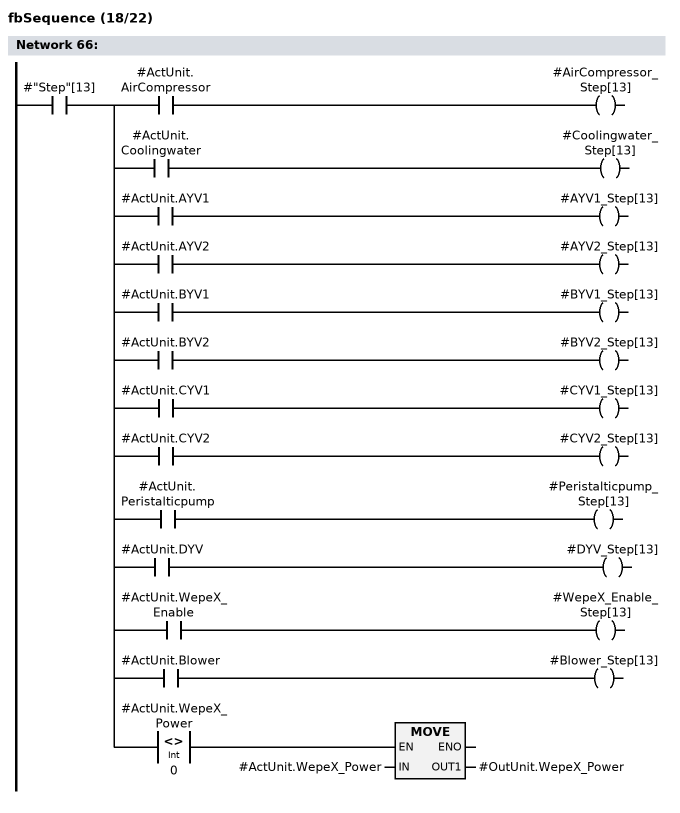
   RUNG wire#powerrail
      Contact( #"Step"[13] )
      wire#w1
      Contact( #ActUnit.AirCompressor )
      Coil( #AirCompressor_Step[13] )
   END_RUNG
   RUNG wire#w1
      Contact( #ActUnit.Coolingwater )
      Coil( #Coolingwater_Step[13] )
   END_RUNG
   RUNG wire#w1
      Contact( #ActUnit.AYV1 )
      Coil( #AYV1_Step[13] )
   END_RUNG
   RUNG wire#w1
      Contact( #ActUnit.AYV2 )
      Coil( #AYV2_Step[13] )
   END_RUNG
   RUNG wire#w1
      Contact( #ActUnit.BYV1 )
      Coil( #BYV1_Step[13] )
   END_RUNG
   RUNG wire#w1
      Contact( #ActUnit.BYV2 )
      Coil( #BYV2_Step[13] )
   END_RUNG
   RUNG wire#w1
      Contact( #ActUnit.CYV1 )
      Coil( #CYV1_Step[13] )
   END_RUNG
   RUNG wire#w1
      Contact( #ActUnit.CYV2 )
      Coil( #CYV2_Step[13] )
   END_RUNG
   RUNG wire#w1
      Contact( #ActUnit.Peristalticpump )
      Coil( #Peristalticpump_Step[13] )
   END_RUNG
   RUNG wire#w1
      Contact( #ActUnit.DYV )
      Coil( #DYV_Step[13] )
   END_RUNG
   RUNG wire#w1
      Contact( #ActUnit.WepeX_Enable )
      Coil( #WepeX_Enable_Step[13] )
   END_RUNG
   RUNG wire#w1
      Contact( #ActUnit.Blower )
      Coil( #Blower_Step[13] )
   END_RUNG
   RUNG wire#w1
      { S7_Templates := "SrcType := Int" } NE_Contact(in1 := #ActUnit.WepeX_Power, in2 := 0)
      Move(in := #ActUnit.WepeX_Power, out1 => #OutUnit.WepeX_Power)
   END_RUNG
   // the same network as SCL:
   #AirCompressor_Step[13] := #"Step"[13] AND #ActUnit.AirCompressor;
   #Coolingwater_Step[13] := #"Step"[13] AND #ActUnit.Coolingwater;
   #AYV1_Step[13] := #"Step"[13] AND #ActUnit.AYV1;
   #AYV2_Step[13] := #"Step"[13] AND #ActUnit.AYV2;
   #BYV1_Step[13] := #"Step"[13] AND #ActUnit.BYV1;
   #BYV2_Step[13] := #"Step"[13] AND #ActUnit.BYV2;
   #CYV1_Step[13] := #"Step"[13] AND #ActUnit.CYV1;
   #CYV2_Step[13] := #"Step"[13] AND #ActUnit.CYV2;
   #Peristalticpump_Step[13] := #"Step"[13] AND #ActUnit.Peristalticpump;
   #DYV_Step[13] := #"Step"[13] AND #ActUnit.DYV;
   #WepeX_Enable_Step[13] := #"Step"[13] AND #ActUnit.WepeX_Enable;
   #Blower_Step[13] := #"Step"[13] AND #ActUnit.Blower;
   IF #"Step"[13] AND (#ActUnit.WepeX_Power <> 0) THEN #OutUnit.WepeX_Power := #ActUnit.WepeX_Power; END_IF;
END_REGION

REGION Network 67
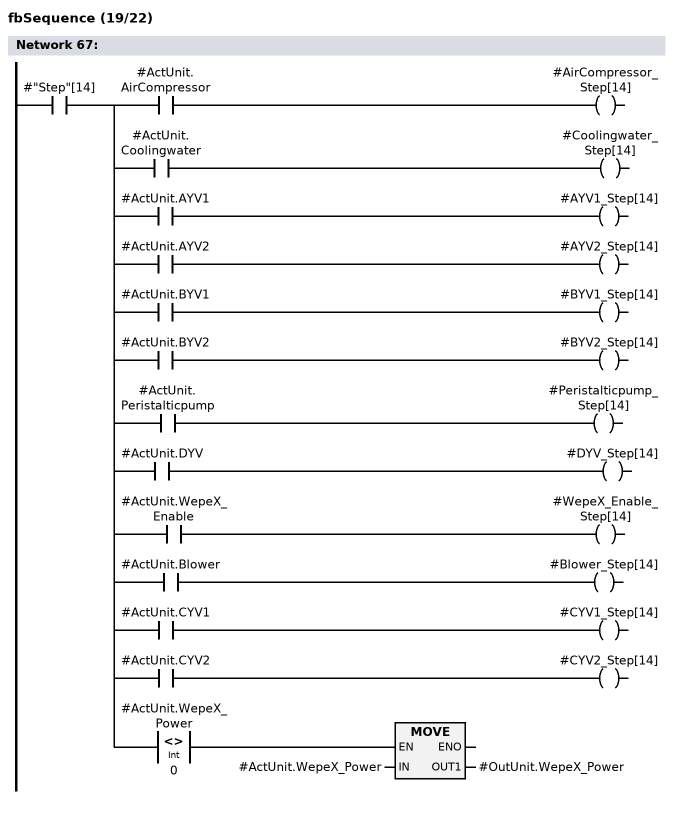
   RUNG wire#powerrail
      Contact( #"Step"[14] )
      wire#w1
      Contact( #ActUnit.AirCompressor )
      Coil( #AirCompressor_Step[14] )
   END_RUNG
   RUNG wire#w1
      Contact( #ActUnit.Coolingwater )
      Coil( #Coolingwater_Step[14] )
   END_RUNG
   RUNG wire#w1
      Contact( #ActUnit.AYV1 )
      Coil( #AYV1_Step[14] )
   END_RUNG
   RUNG wire#w1
      Contact( #ActUnit.AYV2 )
      Coil( #AYV2_Step[14] )
   END_RUNG
   RUNG wire#w1
      Contact( #ActUnit.BYV1 )
      Coil( #BYV1_Step[14] )
   END_RUNG
   RUNG wire#w1
      Contact( #ActUnit.BYV2 )
      Coil( #BYV2_Step[14] )
   END_RUNG
   RUNG wire#w1
      Contact( #ActUnit.Peristalticpump )
      Coil( #Peristalticpump_Step[14] )
   END_RUNG
   RUNG wire#w1
      Contact( #ActUnit.DYV )
      Coil( #DYV_Step[14] )
   END_RUNG
   RUNG wire#w1
      Contact( #ActUnit.WepeX_Enable )
      Coil( #WepeX_Enable_Step[14] )
   END_RUNG
   RUNG wire#w1
      Contact( #ActUnit.Blower )
      Coil( #Blower_Step[14] )
   END_RUNG
   RUNG wire#w1
      Contact( #ActUnit.CYV1 )
      Coil( #CYV1_Step[14] )
   END_RUNG
   RUNG wire#w1
      Contact( #ActUnit.CYV2 )
      Coil( #CYV2_Step[14] )
   END_RUNG
   RUNG wire#w1
      { S7_Templates := "SrcType := Int" } NE_Contact(in1 := #ActUnit.WepeX_Power, in2 := 0)
      Move(in := #ActUnit.WepeX_Power, out1 => #OutUnit.WepeX_Power)
   END_RUNG
   // the same network as SCL:
   #AirCompressor_Step[14] := #"Step"[14] AND #ActUnit.AirCompressor;
   #Coolingwater_Step[14] := #"Step"[14] AND #ActUnit.Coolingwater;
   #AYV1_Step[14] := #"Step"[14] AND #ActUnit.AYV1;
   #AYV2_Step[14] := #"Step"[14] AND #ActUnit.AYV2;
   #BYV1_Step[14] := #"Step"[14] AND #ActUnit.BYV1;
   #BYV2_Step[14] := #"Step"[14] AND #ActUnit.BYV2;
   #Peristalticpump_Step[14] := #"Step"[14] AND #ActUnit.Peristalticpump;
   #DYV_Step[14] := #"Step"[14] AND #ActUnit.DYV;
   #WepeX_Enable_Step[14] := #"Step"[14] AND #ActUnit.WepeX_Enable;
   #Blower_Step[14] := #"Step"[14] AND #ActUnit.Blower;
   #CYV1_Step[14] := #"Step"[14] AND #ActUnit.CYV1;
   #CYV2_Step[14] := #"Step"[14] AND #ActUnit.CYV2;
   IF #"Step"[14] AND (#ActUnit.WepeX_Power <> 0) THEN #OutUnit.WepeX_Power := #ActUnit.WepeX_Power; END_IF;
END_REGION

REGION Network 68
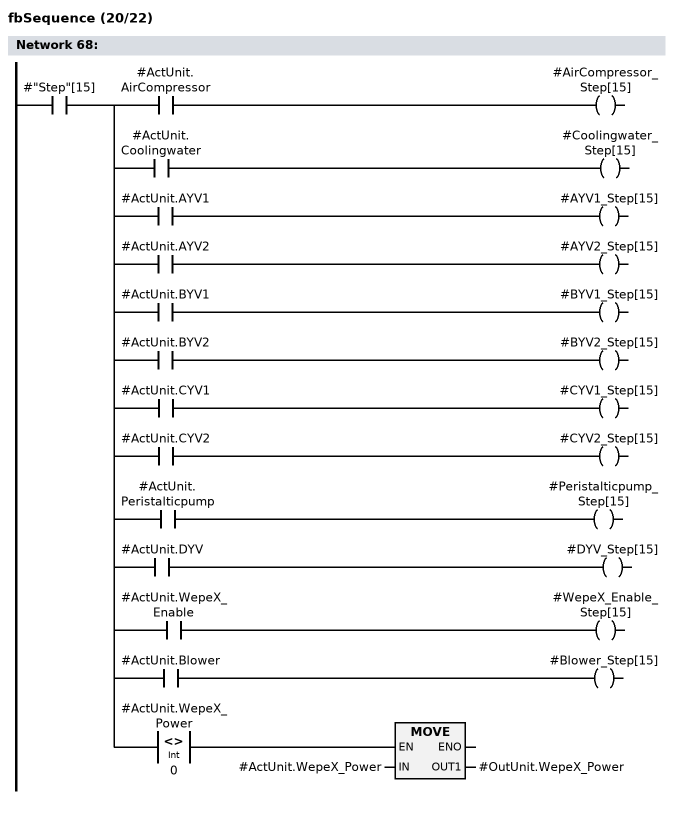
   RUNG wire#powerrail
      Contact( #"Step"[15] )
      wire#w1
      Contact( #ActUnit.AirCompressor )
      Coil( #AirCompressor_Step[15] )
   END_RUNG
   RUNG wire#w1
      Contact( #ActUnit.Coolingwater )
      Coil( #Coolingwater_Step[15] )
   END_RUNG
   RUNG wire#w1
      Contact( #ActUnit.AYV1 )
      Coil( #AYV1_Step[15] )
   END_RUNG
   RUNG wire#w1
      Contact( #ActUnit.AYV2 )
      Coil( #AYV2_Step[15] )
   END_RUNG
   RUNG wire#w1
      Contact( #ActUnit.BYV1 )
      Coil( #BYV1_Step[15] )
   END_RUNG
   RUNG wire#w1
      Contact( #ActUnit.BYV2 )
      Coil( #BYV2_Step[15] )
   END_RUNG
   RUNG wire#w1
      Contact( #ActUnit.CYV1 )
      Coil( #CYV1_Step[15] )
   END_RUNG
   RUNG wire#w1
      Contact( #ActUnit.CYV2 )
      Coil( #CYV2_Step[15] )
   END_RUNG
   RUNG wire#w1
      Contact( #ActUnit.Peristalticpump )
      Coil( #Peristalticpump_Step[15] )
   END_RUNG
   RUNG wire#w1
      Contact( #ActUnit.DYV )
      Coil( #DYV_Step[15] )
   END_RUNG
   RUNG wire#w1
      Contact( #ActUnit.WepeX_Enable )
      Coil( #WepeX_Enable_Step[15] )
   END_RUNG
   RUNG wire#w1
      Contact( #ActUnit.Blower )
      Coil( #Blower_Step[15] )
   END_RUNG
   RUNG wire#w1
      { S7_Templates := "SrcType := Int" } NE_Contact(in1 := #ActUnit.WepeX_Power, in2 := 0)
      Move(in := #ActUnit.WepeX_Power, out1 => #OutUnit.WepeX_Power)
   END_RUNG
   // the same network as SCL:
   #AirCompressor_Step[15] := #"Step"[15] AND #ActUnit.AirCompressor;
   #Coolingwater_Step[15] := #"Step"[15] AND #ActUnit.Coolingwater;
   #AYV1_Step[15] := #"Step"[15] AND #ActUnit.AYV1;
   #AYV2_Step[15] := #"Step"[15] AND #ActUnit.AYV2;
   #BYV1_Step[15] := #"Step"[15] AND #ActUnit.BYV1;
   #BYV2_Step[15] := #"Step"[15] AND #ActUnit.BYV2;
   #CYV1_Step[15] := #"Step"[15] AND #ActUnit.CYV1;
   #CYV2_Step[15] := #"Step"[15] AND #ActUnit.CYV2;
   #Peristalticpump_Step[15] := #"Step"[15] AND #ActUnit.Peristalticpump;
   #DYV_Step[15] := #"Step"[15] AND #ActUnit.DYV;
   #WepeX_Enable_Step[15] := #"Step"[15] AND #ActUnit.WepeX_Enable;
   #Blower_Step[15] := #"Step"[15] AND #ActUnit.Blower;
   IF #"Step"[15] AND (#ActUnit.WepeX_Power <> 0) THEN #OutUnit.WepeX_Power := #ActUnit.WepeX_Power; END_IF;
END_REGION

REGION Network 69
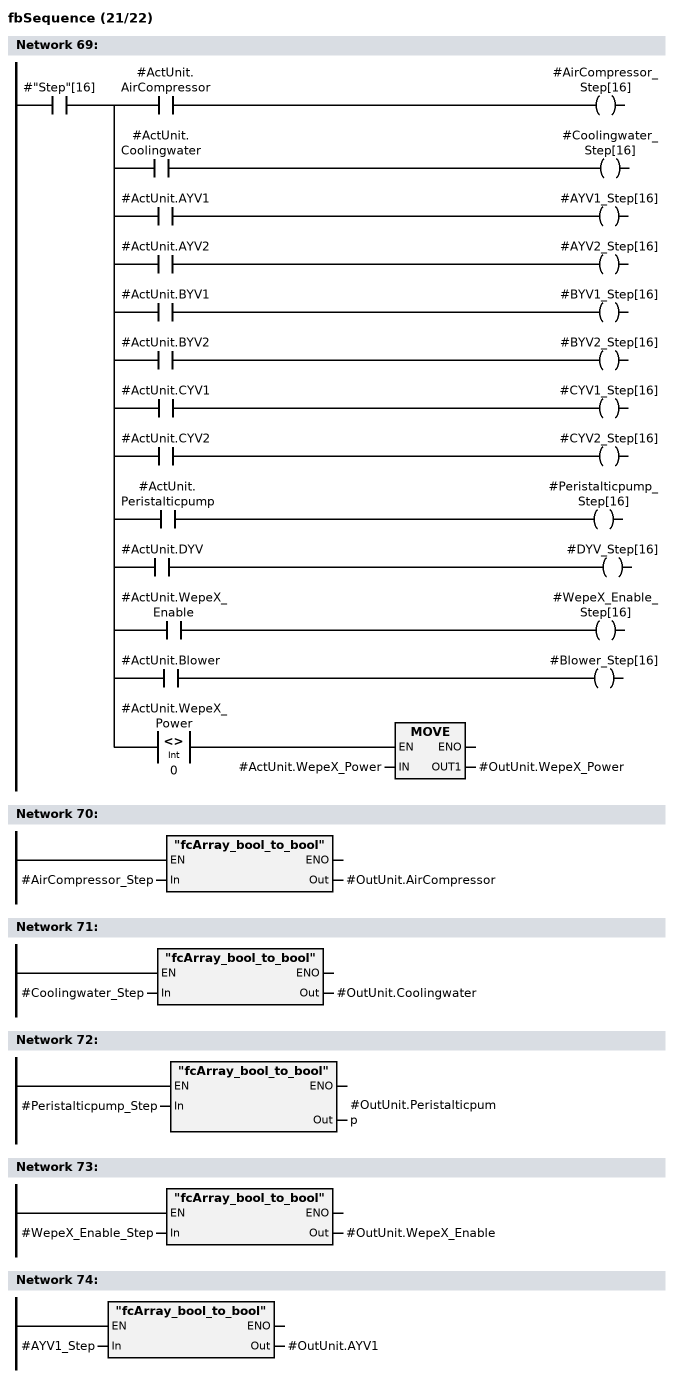
   RUNG wire#powerrail
      Contact( #"Step"[16] )
      wire#w1
      Contact( #ActUnit.AirCompressor )
      Coil( #AirCompressor_Step[16] )
   END_RUNG
   RUNG wire#w1
      Contact( #ActUnit.Coolingwater )
      Coil( #Coolingwater_Step[16] )
   END_RUNG
   RUNG wire#w1
      Contact( #ActUnit.AYV1 )
      Coil( #AYV1_Step[16] )
   END_RUNG
   RUNG wire#w1
      Contact( #ActUnit.AYV2 )
      Coil( #AYV2_Step[16] )
   END_RUNG
   RUNG wire#w1
      Contact( #ActUnit.BYV1 )
      Coil( #BYV1_Step[16] )
   END_RUNG
   RUNG wire#w1
      Contact( #ActUnit.BYV2 )
      Coil( #BYV2_Step[16] )
   END_RUNG
   RUNG wire#w1
      Contact( #ActUnit.CYV1 )
      Coil( #CYV1_Step[16] )
   END_RUNG
   RUNG wire#w1
      Contact( #ActUnit.CYV2 )
      Coil( #CYV2_Step[16] )
   END_RUNG
   RUNG wire#w1
      Contact( #ActUnit.Peristalticpump )
      Coil( #Peristalticpump_Step[16] )
   END_RUNG
   RUNG wire#w1
      Contact( #ActUnit.DYV )
      Coil( #DYV_Step[16] )
   END_RUNG
   RUNG wire#w1
      Contact( #ActUnit.WepeX_Enable )
      Coil( #WepeX_Enable_Step[16] )
   END_RUNG
   RUNG wire#w1
      Contact( #ActUnit.Blower )
      Coil( #Blower_Step[16] )
   END_RUNG
   RUNG wire#w1
      { S7_Templates := "SrcType := Int" } NE_Contact(in1 := #ActUnit.WepeX_Power, in2 := 0)
      Move(in := #ActUnit.WepeX_Power, out1 => #OutUnit.WepeX_Power)
   END_RUNG
   // the same network as SCL:
   #AirCompressor_Step[16] := #"Step"[16] AND #ActUnit.AirCompressor;
   #Coolingwater_Step[16] := #"Step"[16] AND #ActUnit.Coolingwater;
   #AYV1_Step[16] := #"Step"[16] AND #ActUnit.AYV1;
   #AYV2_Step[16] := #"Step"[16] AND #ActUnit.AYV2;
   #BYV1_Step[16] := #"Step"[16] AND #ActUnit.BYV1;
   #BYV2_Step[16] := #"Step"[16] AND #ActUnit.BYV2;
   #CYV1_Step[16] := #"Step"[16] AND #ActUnit.CYV1;
   #CYV2_Step[16] := #"Step"[16] AND #ActUnit.CYV2;
   #Peristalticpump_Step[16] := #"Step"[16] AND #ActUnit.Peristalticpump;
   #DYV_Step[16] := #"Step"[16] AND #ActUnit.DYV;
   #WepeX_Enable_Step[16] := #"Step"[16] AND #ActUnit.WepeX_Enable;
   #Blower_Step[16] := #"Step"[16] AND #ActUnit.Blower;
   IF #"Step"[16] AND (#ActUnit.WepeX_Power <> 0) THEN #OutUnit.WepeX_Power := #ActUnit.WepeX_Power; END_IF;
END_REGION

REGION Network 70
   RUNG wire#powerrail
      "fcArray_bool_to_bool"(In := #AirCompressor_Step, Out => #OutUnit.AirCompressor)
   END_RUNG
   // the same network as SCL:
   "fcArray_bool_to_bool"(In := #AirCompressor_Step, Out => #OutUnit.AirCompressor);
END_REGION

REGION Network 71
   RUNG wire#powerrail
      "fcArray_bool_to_bool"(In := #Coolingwater_Step, Out => #OutUnit.Coolingwater)
   END_RUNG
   // the same network as SCL:
   "fcArray_bool_to_bool"(In := #Coolingwater_Step, Out => #OutUnit.Coolingwater);
END_REGION

REGION Network 72
   RUNG wire#powerrail
      "fcArray_bool_to_bool"(In := #Peristalticpump_Step, Out => #OutUnit.Peristalticpump)
   END_RUNG
   // the same network as SCL:
   "fcArray_bool_to_bool"(In := #Peristalticpump_Step, Out => #OutUnit.Peristalticpump);
END_REGION

REGION Network 73
   RUNG wire#powerrail
      "fcArray_bool_to_bool"(In := #WepeX_Enable_Step, Out => #OutUnit.WepeX_Enable)
   END_RUNG
   // the same network as SCL:
   "fcArray_bool_to_bool"(In := #WepeX_Enable_Step, Out => #OutUnit.WepeX_Enable);
END_REGION

REGION Network 74
   RUNG wire#powerrail
      "fcArray_bool_to_bool"(In := #AYV1_Step, Out => #OutUnit.AYV1)
   END_RUNG
   // the same network as SCL:
   "fcArray_bool_to_bool"(In := #AYV1_Step, Out => #OutUnit.AYV1);
END_REGION

REGION Network 75
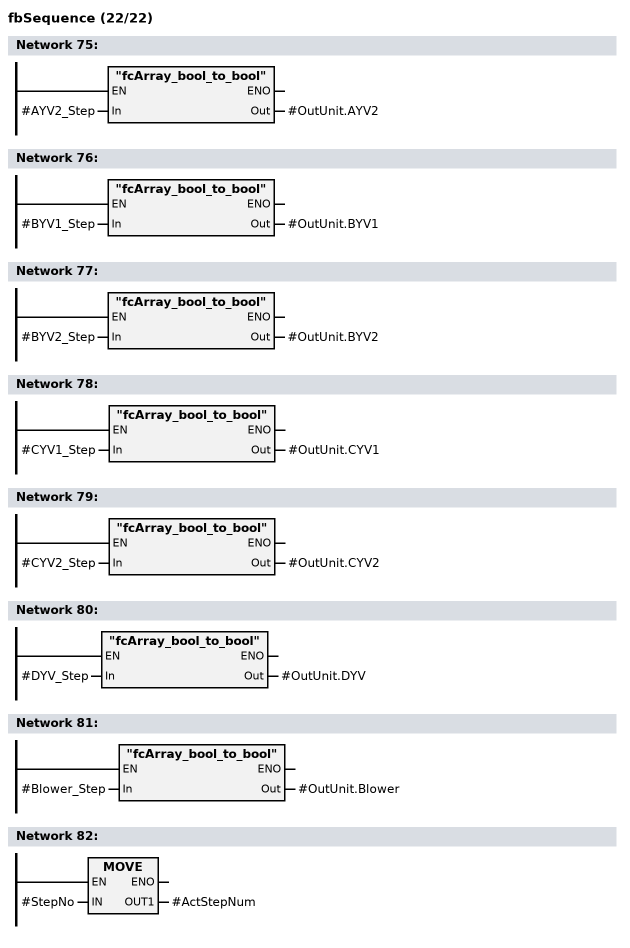
   RUNG wire#powerrail
      "fcArray_bool_to_bool"(In := #AYV2_Step, Out => #OutUnit.AYV2)
   END_RUNG
   // the same network as SCL:
   "fcArray_bool_to_bool"(In := #AYV2_Step, Out => #OutUnit.AYV2);
END_REGION

REGION Network 76
   RUNG wire#powerrail
      "fcArray_bool_to_bool"(In := #BYV1_Step, Out => #OutUnit.BYV1)
   END_RUNG
   // the same network as SCL:
   "fcArray_bool_to_bool"(In := #BYV1_Step, Out => #OutUnit.BYV1);
END_REGION

REGION Network 77
   RUNG wire#powerrail
      "fcArray_bool_to_bool"(In := #BYV2_Step, Out => #OutUnit.BYV2)
   END_RUNG
   // the same network as SCL:
   "fcArray_bool_to_bool"(In := #BYV2_Step, Out => #OutUnit.BYV2);
END_REGION

REGION Network 78
   RUNG wire#powerrail
      "fcArray_bool_to_bool"(In := #CYV1_Step, Out => #OutUnit.CYV1)
   END_RUNG
   // the same network as SCL:
   "fcArray_bool_to_bool"(In := #CYV1_Step, Out => #OutUnit.CYV1);
END_REGION

REGION Network 79
   RUNG wire#powerrail
      "fcArray_bool_to_bool"(In := #CYV2_Step, Out => #OutUnit.CYV2)
   END_RUNG
   // the same network as SCL:
   "fcArray_bool_to_bool"(In := #CYV2_Step, Out => #OutUnit.CYV2);
END_REGION

REGION Network 80
   RUNG wire#powerrail
      "fcArray_bool_to_bool"(In := #DYV_Step, Out => #OutUnit.DYV)
   END_RUNG
   // the same network as SCL:
   "fcArray_bool_to_bool"(In := #DYV_Step, Out => #OutUnit.DYV);
END_REGION

REGION Network 81
   RUNG wire#powerrail
      "fcArray_bool_to_bool"(In := #Blower_Step, Out => #OutUnit.Blower)
   END_RUNG
   // the same network as SCL:
   "fcArray_bool_to_bool"(In := #Blower_Step, Out => #OutUnit.Blower);
END_REGION

REGION Network 82
   RUNG wire#powerrail
      Move(in := #StepNo, out1 => #ActStepNum)
   END_RUNG
   // the same network as SCL:
   #ActStepNum := #StepNo;
END_REGION
END_FUNCTION_BLOCK

FUNCTION "fcDataMv" : Void   // FC100, LAD
{ S7_Optimized_Access := 'TRUE' }
VERSION : 0.1
BEGIN

REGION Network 1
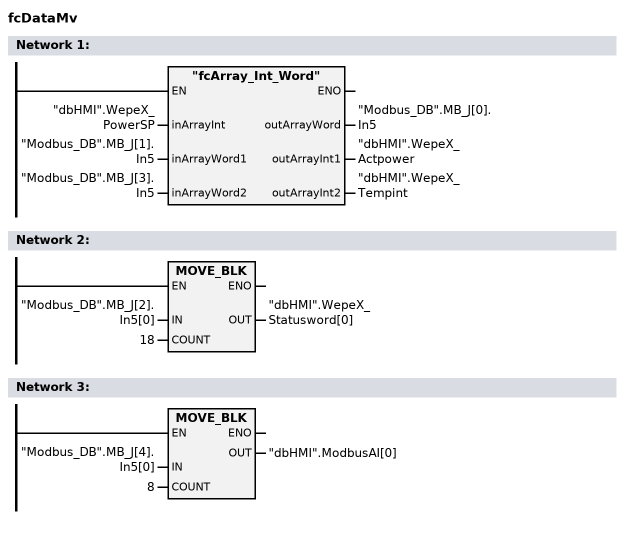
   RUNG wire#powerrail
      "fcArray_Int_Word"(inArrayInt := "dbHMI".WepeX_PowerSP, inArrayWord1 := "Modbus_DB".MB_J[1].In5, inArrayWord2 := "Modbus_DB".MB_J[3].In5, outArrayWord => "Modbus_DB".MB_J[0].In5, outArrayInt1 => "dbHMI".WepeX_Actpower, outArrayInt2 => "dbHMI".WepeX_Tempint)
   END_RUNG
   // the same network as SCL:
   "fcArray_Int_Word"(inArrayInt := "dbHMI".WepeX_PowerSP,
                      inArrayWord1 := "Modbus_DB".MB_J[1].In5,
                      inArrayWord2 := "Modbus_DB".MB_J[3].In5,
                      outArrayWord => "Modbus_DB".MB_J[0].In5,
                      outArrayInt1 => "dbHMI".WepeX_Actpower,
                      outArrayInt2 => "dbHMI".WepeX_Tempint);
END_REGION

REGION Network 2
   MOVE_BLK(IN := "Modbus_DB".MB_J[2].In5[0], COUNT := 18, OUT => "dbHMI".WepeX_Statusword[0]);
END_REGION

REGION Network 3
   MOVE_BLK(IN := "Modbus_DB".MB_J[4].In5[0], COUNT := 8, OUT => "dbHMI".ModbusAI[0]);
END_REGION
END_FUNCTION

FUNCTION "fcArray_Int_Word" : Void   // FC101, LAD
{ S7_Optimized_Access := 'TRUE' }
VERSION : 0.1
   VAR_INPUT
      inArrayInt : Array[0..17] of Int;
      inArrayWord1 : Array[0..17] of Word;
      inArrayWord2 : Array[0..17] of Word;
   END_VAR
   VAR_OUTPUT
      outArrayWord : Array[0..17] of Word;
      outArrayInt1 : Array[0..17] of Int;
      outArrayInt2 : Array[0..17] of Int;
   END_VAR
BEGIN

REGION Network 1
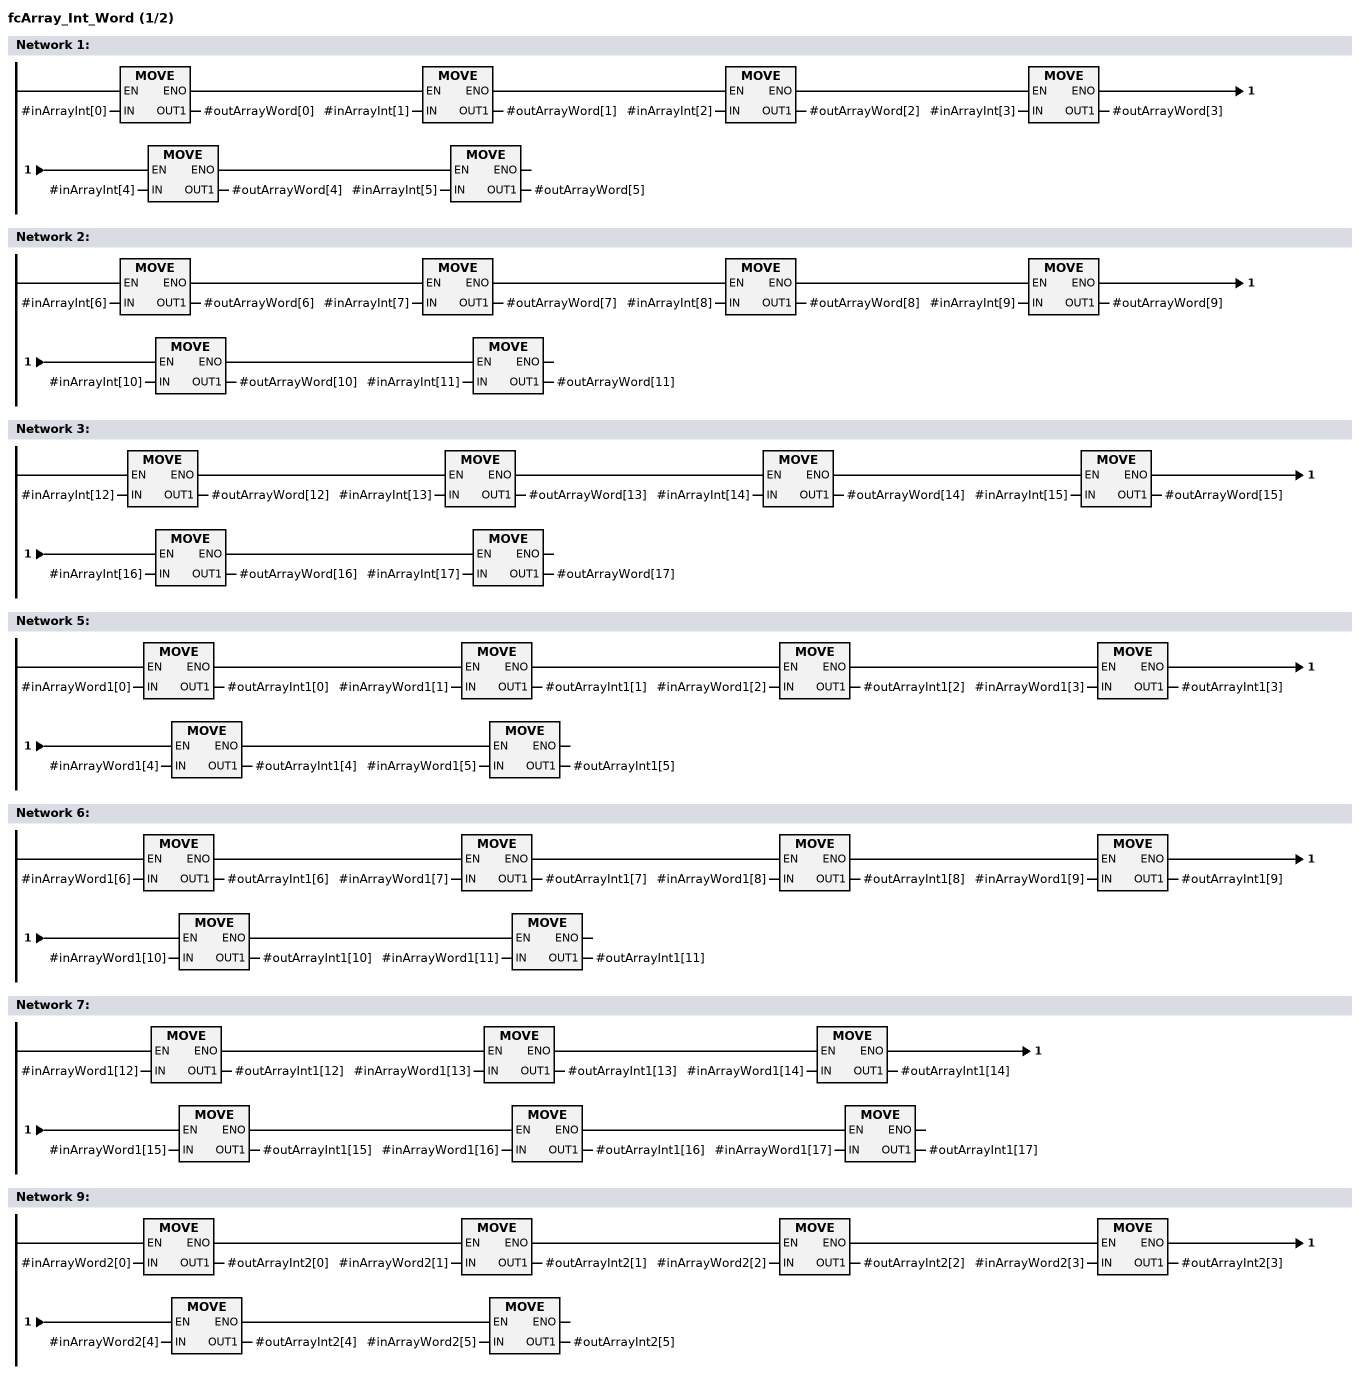
   RUNG wire#powerrail
      Move(in := #inArrayInt[0], out1 => #outArrayWord[0])
      Move(in := #inArrayInt[1], out1 => #outArrayWord[1])
      Move(in := #inArrayInt[2], out1 => #outArrayWord[2])
      Move(in := #inArrayInt[3], out1 => #outArrayWord[3])
      Move(in := #inArrayInt[4], out1 => #outArrayWord[4])
      Move(in := #inArrayInt[5], out1 => #outArrayWord[5])
   END_RUNG
   // the same network as SCL:
   #outArrayWord[0] := #inArrayInt[0];
   #outArrayWord[1] := #inArrayInt[1];
   #outArrayWord[2] := #inArrayInt[2];
   #outArrayWord[3] := #inArrayInt[3];
   #outArrayWord[4] := #inArrayInt[4];
   #outArrayWord[5] := #inArrayInt[5];
END_REGION

REGION Network 2
   RUNG wire#powerrail
      Move(in := #inArrayInt[6], out1 => #outArrayWord[6])
      Move(in := #inArrayInt[7], out1 => #outArrayWord[7])
      Move(in := #inArrayInt[8], out1 => #outArrayWord[8])
      Move(in := #inArrayInt[9], out1 => #outArrayWord[9])
      Move(in := #inArrayInt[10], out1 => #outArrayWord[10])
      Move(in := #inArrayInt[11], out1 => #outArrayWord[11])
   END_RUNG
   // the same network as SCL:
   #outArrayWord[6] := #inArrayInt[6];
   #outArrayWord[7] := #inArrayInt[7];
   #outArrayWord[8] := #inArrayInt[8];
   #outArrayWord[9] := #inArrayInt[9];
   #outArrayWord[10] := #inArrayInt[10];
   #outArrayWord[11] := #inArrayInt[11];
END_REGION

REGION Network 3
   RUNG wire#powerrail
      Move(in := #inArrayInt[12], out1 => #outArrayWord[12])
      Move(in := #inArrayInt[13], out1 => #outArrayWord[13])
      Move(in := #inArrayInt[14], out1 => #outArrayWord[14])
      Move(in := #inArrayInt[15], out1 => #outArrayWord[15])
      Move(in := #inArrayInt[16], out1 => #outArrayWord[16])
      Move(in := #inArrayInt[17], out1 => #outArrayWord[17])
   END_RUNG
   // the same network as SCL:
   #outArrayWord[12] := #inArrayInt[12];
   #outArrayWord[13] := #inArrayInt[13];
   #outArrayWord[14] := #inArrayInt[14];
   #outArrayWord[15] := #inArrayInt[15];
   #outArrayWord[16] := #inArrayInt[16];
   #outArrayWord[17] := #inArrayInt[17];
END_REGION

REGION Network 5
   RUNG wire#powerrail
      Move(in := #inArrayWord1[0], out1 => #outArrayInt1[0])
      Move(in := #inArrayWord1[1], out1 => #outArrayInt1[1])
      Move(in := #inArrayWord1[2], out1 => #outArrayInt1[2])
      Move(in := #inArrayWord1[3], out1 => #outArrayInt1[3])
      Move(in := #inArrayWord1[4], out1 => #outArrayInt1[4])
      Move(in := #inArrayWord1[5], out1 => #outArrayInt1[5])
   END_RUNG
   // the same network as SCL:
   #outArrayInt1[0] := #inArrayWord1[0];
   #outArrayInt1[1] := #inArrayWord1[1];
   #outArrayInt1[2] := #inArrayWord1[2];
   #outArrayInt1[3] := #inArrayWord1[3];
   #outArrayInt1[4] := #inArrayWord1[4];
   #outArrayInt1[5] := #inArrayWord1[5];
END_REGION

REGION Network 6
   RUNG wire#powerrail
      Move(in := #inArrayWord1[6], out1 => #outArrayInt1[6])
      Move(in := #inArrayWord1[7], out1 => #outArrayInt1[7])
      Move(in := #inArrayWord1[8], out1 => #outArrayInt1[8])
      Move(in := #inArrayWord1[9], out1 => #outArrayInt1[9])
      Move(in := #inArrayWord1[10], out1 => #outArrayInt1[10])
      Move(in := #inArrayWord1[11], out1 => #outArrayInt1[11])
   END_RUNG
   // the same network as SCL:
   #outArrayInt1[6] := #inArrayWord1[6];
   #outArrayInt1[7] := #inArrayWord1[7];
   #outArrayInt1[8] := #inArrayWord1[8];
   #outArrayInt1[9] := #inArrayWord1[9];
   #outArrayInt1[10] := #inArrayWord1[10];
   #outArrayInt1[11] := #inArrayWord1[11];
END_REGION

REGION Network 7
   RUNG wire#powerrail
      Move(in := #inArrayWord1[12], out1 => #outArrayInt1[12])
      Move(in := #inArrayWord1[13], out1 => #outArrayInt1[13])
      Move(in := #inArrayWord1[14], out1 => #outArrayInt1[14])
      Move(in := #inArrayWord1[15], out1 => #outArrayInt1[15])
      Move(in := #inArrayWord1[16], out1 => #outArrayInt1[16])
      Move(in := #inArrayWord1[17], out1 => #outArrayInt1[17])
   END_RUNG
   // the same network as SCL:
   #outArrayInt1[12] := #inArrayWord1[12];
   #outArrayInt1[13] := #inArrayWord1[13];
   #outArrayInt1[14] := #inArrayWord1[14];
   #outArrayInt1[15] := #inArrayWord1[15];
   #outArrayInt1[16] := #inArrayWord1[16];
   #outArrayInt1[17] := #inArrayWord1[17];
END_REGION

REGION Network 9
   RUNG wire#powerrail
      Move(in := #inArrayWord2[0], out1 => #outArrayInt2[0])
      Move(in := #inArrayWord2[1], out1 => #outArrayInt2[1])
      Move(in := #inArrayWord2[2], out1 => #outArrayInt2[2])
      Move(in := #inArrayWord2[3], out1 => #outArrayInt2[3])
      Move(in := #inArrayWord2[4], out1 => #outArrayInt2[4])
      Move(in := #inArrayWord2[5], out1 => #outArrayInt2[5])
   END_RUNG
   // the same network as SCL:
   #outArrayInt2[0] := #inArrayWord2[0];
   #outArrayInt2[1] := #inArrayWord2[1];
   #outArrayInt2[2] := #inArrayWord2[2];
   #outArrayInt2[3] := #inArrayWord2[3];
   #outArrayInt2[4] := #inArrayWord2[4];
   #outArrayInt2[5] := #inArrayWord2[5];
END_REGION

REGION Network 10
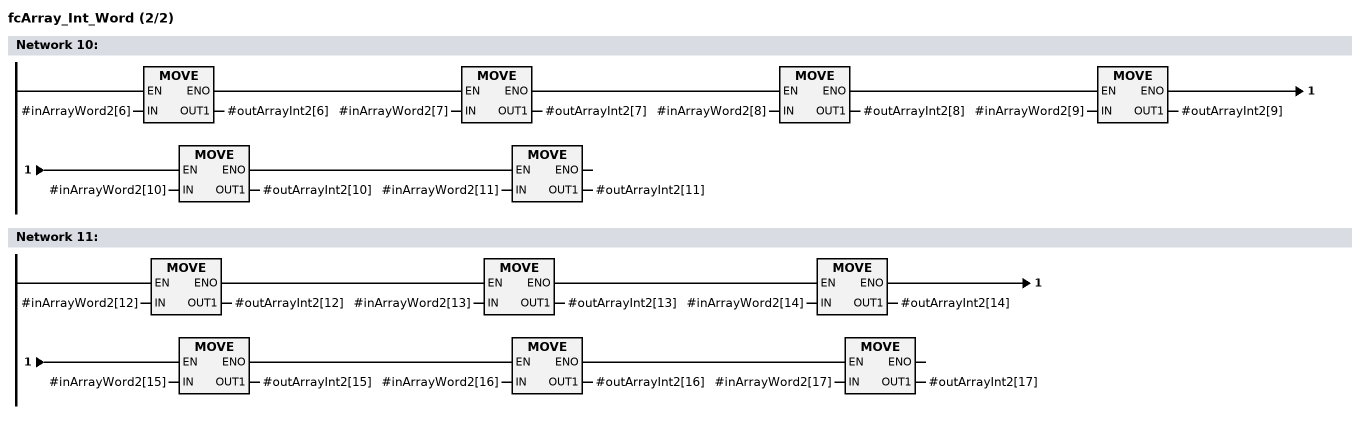
   RUNG wire#powerrail
      Move(in := #inArrayWord2[6], out1 => #outArrayInt2[6])
      Move(in := #inArrayWord2[7], out1 => #outArrayInt2[7])
      Move(in := #inArrayWord2[8], out1 => #outArrayInt2[8])
      Move(in := #inArrayWord2[9], out1 => #outArrayInt2[9])
      Move(in := #inArrayWord2[10], out1 => #outArrayInt2[10])
      Move(in := #inArrayWord2[11], out1 => #outArrayInt2[11])
   END_RUNG
   // the same network as SCL:
   #outArrayInt2[6] := #inArrayWord2[6];
   #outArrayInt2[7] := #inArrayWord2[7];
   #outArrayInt2[8] := #inArrayWord2[8];
   #outArrayInt2[9] := #inArrayWord2[9];
   #outArrayInt2[10] := #inArrayWord2[10];
   #outArrayInt2[11] := #inArrayWord2[11];
END_REGION

REGION Network 11
   RUNG wire#powerrail
      Move(in := #inArrayWord2[12], out1 => #outArrayInt2[12])
      Move(in := #inArrayWord2[13], out1 => #outArrayInt2[13])
      Move(in := #inArrayWord2[14], out1 => #outArrayInt2[14])
      Move(in := #inArrayWord2[15], out1 => #outArrayInt2[15])
      Move(in := #inArrayWord2[16], out1 => #outArrayInt2[16])
      Move(in := #inArrayWord2[17], out1 => #outArrayInt2[17])
   END_RUNG
   // the same network as SCL:
   #outArrayInt2[12] := #inArrayWord2[12];
   #outArrayInt2[13] := #inArrayWord2[13];
   #outArrayInt2[14] := #inArrayWord2[14];
   #outArrayInt2[15] := #inArrayWord2[15];
   #outArrayInt2[16] := #inArrayWord2[16];
   #outArrayInt2[17] := #inArrayWord2[17];
END_REGION
END_FUNCTION

FUNCTION "fcWepeXStaus" : Void   // FC102, LAD
{ S7_Optimized_Access := 'TRUE' }
VERSION : 0.1
   VAR_INPUT
      Lbyte : Byte;
   END_VAR
   VAR_OUTPUT
      通信不正常 : Bool;
      工作正常 : Bool;
      无反馈信号 : Bool;
      欠压保护 : Bool;
      过压保护 : Bool;
      过流保护 : Bool;
      过温保护 : Bool;
      磁控管故障 : Bool;
      浪涌保护 : Bool;
      高压故障 : Bool;
      开关管故障 : Bool;
      无功率信号 : Bool;
      Vcc保护 : Bool;
      Error : Word;
   END_VAR
BEGIN

REGION Network 1
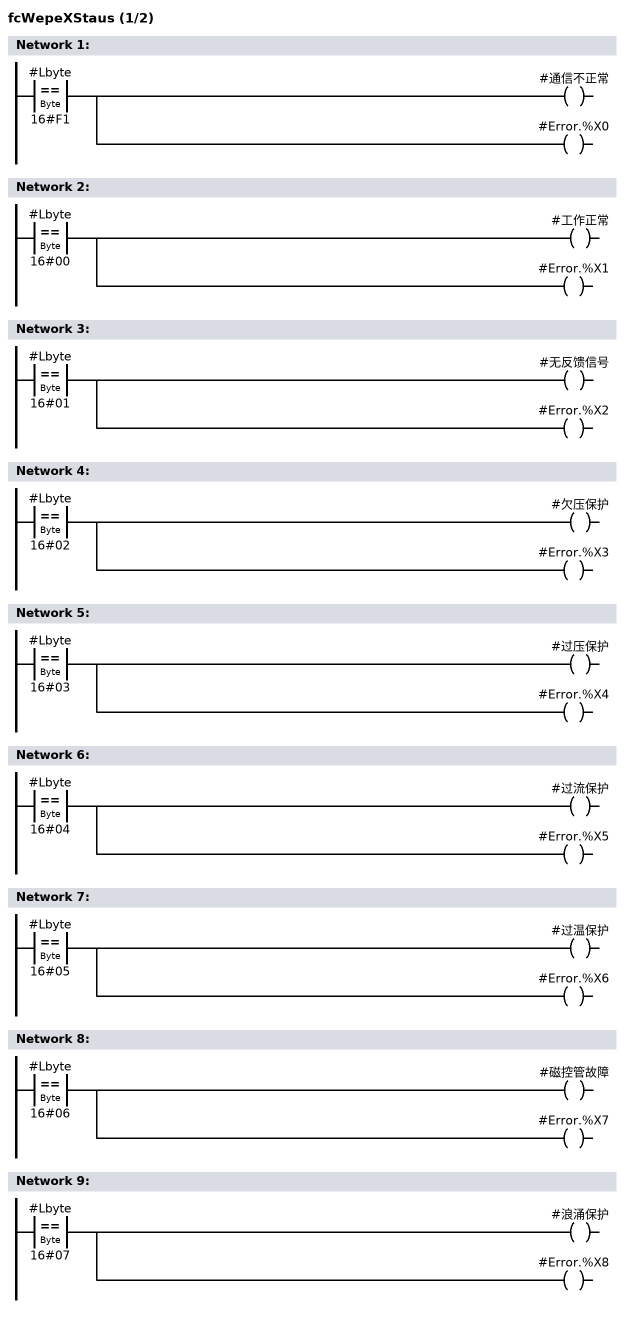
   RUNG wire#powerrail
      { S7_Templates := "SrcType := Byte" } EQ_Contact(in1 := #Lbyte, in2 := 16#F1)
      wire#w1
      Coil( #通信不正常 )
   END_RUNG
   RUNG wire#w1
      Coil( #Error.%X0 )
   END_RUNG
   // the same network as SCL:
   #通信不正常 := #Lbyte = 16#F1;
   #Error.%X0 := #通信不正常;
END_REGION
